
       "Centrifuge_Write_TO_T-103_DB".RequestProduct := "Centrifuge_Write_TO_T-103_DB".RouteOpened AND NOT "Centrifuge_Aux_DB"."Bool".Centrifuge.Status.FeelerRetracted;
       //************************************************Interlocks to T-104*************************************************//
       "Centrifuge_Write_TO_T-104_DB".RouteOpened := "XV-1045_DB".OS AND ("XV-3013_DB".OS OR "XV-3012_DB".OS) AND ("P-301A_DB".CF OR "P-301A_DB".CF);

       "Centrifuge_Write_TO_T-104_DB".ReqWater := "Centrifuge_DB".Status.Step = 29 AND  "Centrifuge_Write_TO_T-104_DB".RouteOpened
       AND NOT "LT-1051_DB".Alarms.HighHigh AND NOT "Centrifuge_DB".Cmds.Hold;
       //***************Valves Status***************//
       "Centrifuge_Aux_DB"."Bool".TOff := "Centrifuge_DB".Equipments.Valves."XV-1045".TurningOff OR "Centrifuge_DB".Equipments.Valves."XV-3013".TurningOff
       OR "Centrifuge_DB".Equipments.Valves."XV-3012".TurningOff OR "Centrifuge_DB".Equipments.Valves."XV-3011".TurningOff;

       //***********************************************Timers****************************************************************************//
       "Centrifuge_Aux_DB"."Bool".WaitForBucketEn := "Centrifuge_DB".Status.Step=26 AND "FT-3011_DB".SAI>1.0;
       "Centrifuge_Aux_DB"."Bool".DryingWetCakeEn := "Centrifuge_DB".Status.Step = 31  AND ("P-301A_DB".CF OR "P-301B_DB".CF) AND "FT-3012_DB".SAI < 0.1; //AND "VFD-C301R_DB".RUN_FEEDBACK
       "Centrifuge_Aux_DB"."Bool".DryingWetCake_Reset := "Centrifuge_DB".Cmds.Abort OR "Centrifuge_DB".Status.Step = 1;
       //Delay for Dry Spin Done to Finish
       "Centrifuge_Aux_DB"."Bool".DrySpinDnDelay_Enab := "Centrifuge_DB".Status.Step = 31 AND "FT-3012_DB".SAI < 0.1 AND ("P-301A_DB".CF OR "P-301B_DB".CF);
END_FUNCTION

FUNCTION "Centrifuge_SEQ_FC" : Void   // FC91, LAD
{ S7_Optimized_Access := 'TRUE' }
VERSION : 0.1
   VAR_TEMP   // added for the SCL form of the ladder/FBD networks
      _w1 : Bool;
      _w2 : Bool;
   END_VAR
BEGIN

REGION Network 2: Abort
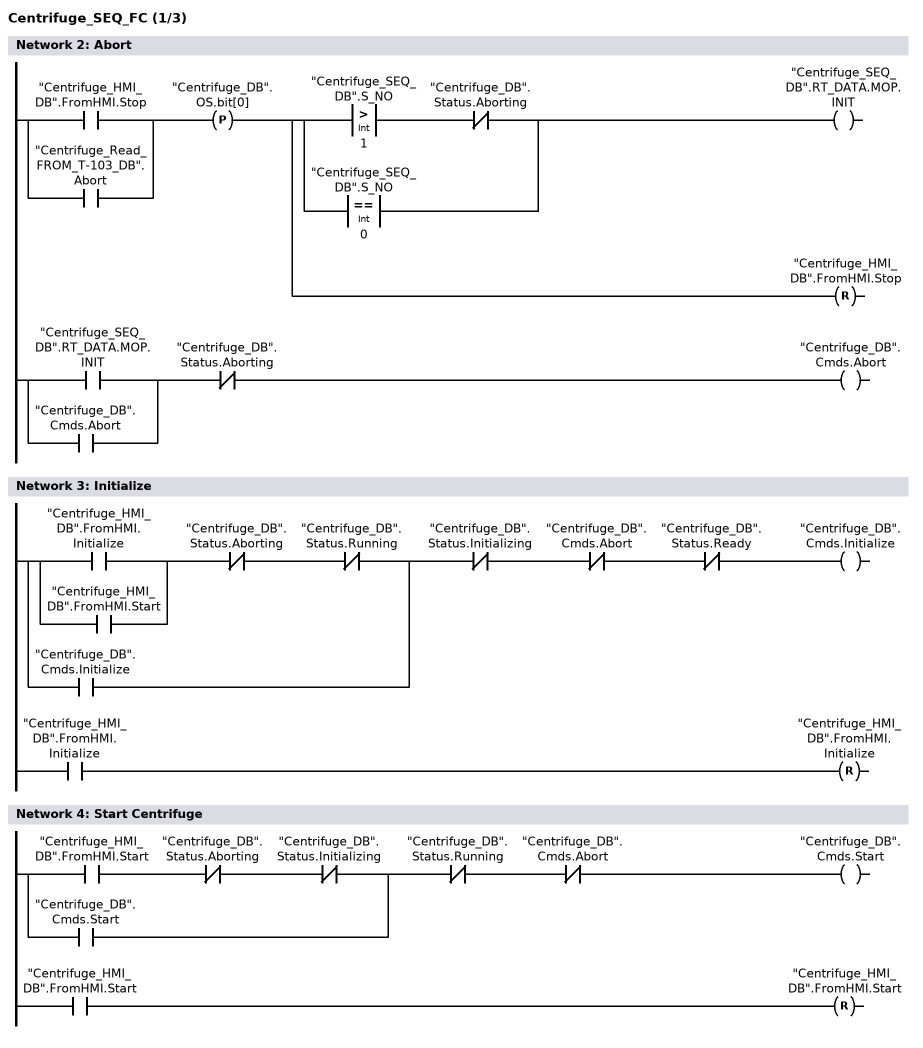
   RUNG wire#powerrail
      Contact( "Centrifuge_HMI_DB".FromHMI.Stop )
      wire#w1
      P_Trig( "Centrifuge_DB".OS.bit[0] )
      wire#w2
      { S7_Templates := "SrcType := Int" } GT_Contact(in1 := "Centrifuge_SEQ_DB".S_NO, in2 := 1)
      I_Contact( "Centrifuge_DB".Status.Aborting )
      wire#w3
      Coil( "Centrifuge_SEQ_DB".RT_DATA.MOP.INIT )
   END_RUNG
   RUNG wire#powerrail
      Contact( "Centrifuge_Read_FROM_T-103_DB".Abort )
   END_RUNG wire#w1
   RUNG wire#w2
      { S7_Templates := "SrcType := Int" } EQ_Contact(in1 := "Centrifuge_SEQ_DB".S_NO, in2 := 0)
   END_RUNG wire#w3
   RUNG wire#w2
      R_Coil( "Centrifuge_HMI_DB".FromHMI.Stop )
   END_RUNG
   RUNG wire#powerrail
      Contact( "Centrifuge_SEQ_DB".RT_DATA.MOP.INIT )
      wire#w4
      I_Contact( "Centrifuge_DB".Status.Aborting )
      Coil( "Centrifuge_DB".Cmds.Abort )
   END_RUNG
   RUNG wire#powerrail
      Contact( "Centrifuge_DB".Cmds.Abort )
   END_RUNG wire#w4
   // the same network as SCL:
   #_w1 := "Centrifuge_HMI_DB".FromHMI.Stop OR "Centrifuge_Read_FROM_T-103_DB".Abort;
   #_w2 := #_w1 AND NOT "Centrifuge_DB".OS.bit[0];   // rising edge
   "Centrifuge_DB".OS.bit[0] := #_w1;
   "Centrifuge_SEQ_DB".RT_DATA.MOP.INIT := #_w2 AND ((("Centrifuge_SEQ_DB".S_NO > 1) AND NOT "Centrifuge_DB".Status.Aborting) OR ("Centrifuge_SEQ_DB".S_NO = 0));
   IF #_w2 THEN "Centrifuge_HMI_DB".FromHMI.Stop := FALSE; END_IF;
   "Centrifuge_DB".Cmds.Abort := ("Centrifuge_SEQ_DB".RT_DATA.MOP.INIT OR "Centrifuge_DB".Cmds.Abort) AND NOT "Centrifuge_DB".Status.Aborting;
END_REGION

REGION Network 3: Initialize
   RUNG wire#powerrail
      Contact( "Centrifuge_HMI_DB".FromHMI.Initialize )
      wire#w1
      I_Contact( "Centrifuge_DB".Status.Aborting )
      I_Contact( "Centrifuge_DB".Status.Running )
      wire#w2
      I_Contact( "Centrifuge_DB".Status.Initializing )
      I_Contact( "Centrifuge_DB".Cmds.Abort )
      I_Contact( "Centrifuge_DB".Status.Ready )
      Coil( "Centrifuge_DB".Cmds.Initialize )
   END_RUNG
   RUNG wire#powerrail
      Contact( "Centrifuge_HMI_DB".FromHMI.Start )
   END_RUNG wire#w1
   RUNG wire#powerrail
      Contact( "Centrifuge_DB".Cmds.Initialize )
   END_RUNG wire#w2
   RUNG wire#powerrail
      Contact( "Centrifuge_HMI_DB".FromHMI.Initialize )
      R_Coil( "Centrifuge_HMI_DB".FromHMI.Initialize )
   END_RUNG
   // the same network as SCL:
   "Centrifuge_DB".Cmds.Initialize := ((("Centrifuge_HMI_DB".FromHMI.Initialize OR "Centrifuge_HMI_DB".FromHMI.Start) AND NOT "Centrifuge_DB".Status.Aborting AND NOT "Centrifuge_DB".Status.Running) OR "Centrifuge_DB".Cmds.Initialize) AND NOT "Centrifuge_DB".Status.Initializing AND NOT "Centrifuge_DB".Cmds.Abort AND NOT "Centrifuge_DB".Status.Ready;
   IF "Centrifuge_HMI_DB".FromHMI.Initialize THEN "Centrifuge_HMI_DB".FromHMI.Initialize := FALSE; END_IF;
END_REGION

REGION Network 4: Start Centrifuge
   RUNG wire#powerrail
      Contact( "Centrifuge_HMI_DB".FromHMI.Start )
      I_Contact( "Centrifuge_DB".Status.Aborting )
      I_Contact( "Centrifuge_DB".Status.Initializing )
      wire#w1
      I_Contact( "Centrifuge_DB".Status.Running )
      I_Contact( "Centrifuge_DB".Cmds.Abort )
      Coil( "Centrifuge_DB".Cmds.Start )
   END_RUNG
   RUNG wire#powerrail
      Contact( "Centrifuge_DB".Cmds.Start )
   END_RUNG wire#w1
   RUNG wire#powerrail
      Contact( "Centrifuge_HMI_DB".FromHMI.Start )
      R_Coil( "Centrifuge_HMI_DB".FromHMI.Start )
   END_RUNG
   // the same network as SCL:
   "Centrifuge_DB".Cmds.Start := (("Centrifuge_HMI_DB".FromHMI.Start AND NOT "Centrifuge_DB".Status.Aborting AND NOT "Centrifuge_DB".Status.Initializing) OR "Centrifuge_DB".Cmds.Start) AND NOT "Centrifuge_DB".Status.Running AND NOT "Centrifuge_DB".Cmds.Abort;
   IF "Centrifuge_HMI_DB".FromHMI.Start THEN "Centrifuge_HMI_DB".FromHMI.Start := FALSE; END_IF;
END_REGION

REGION Network 5: Procedure Selected
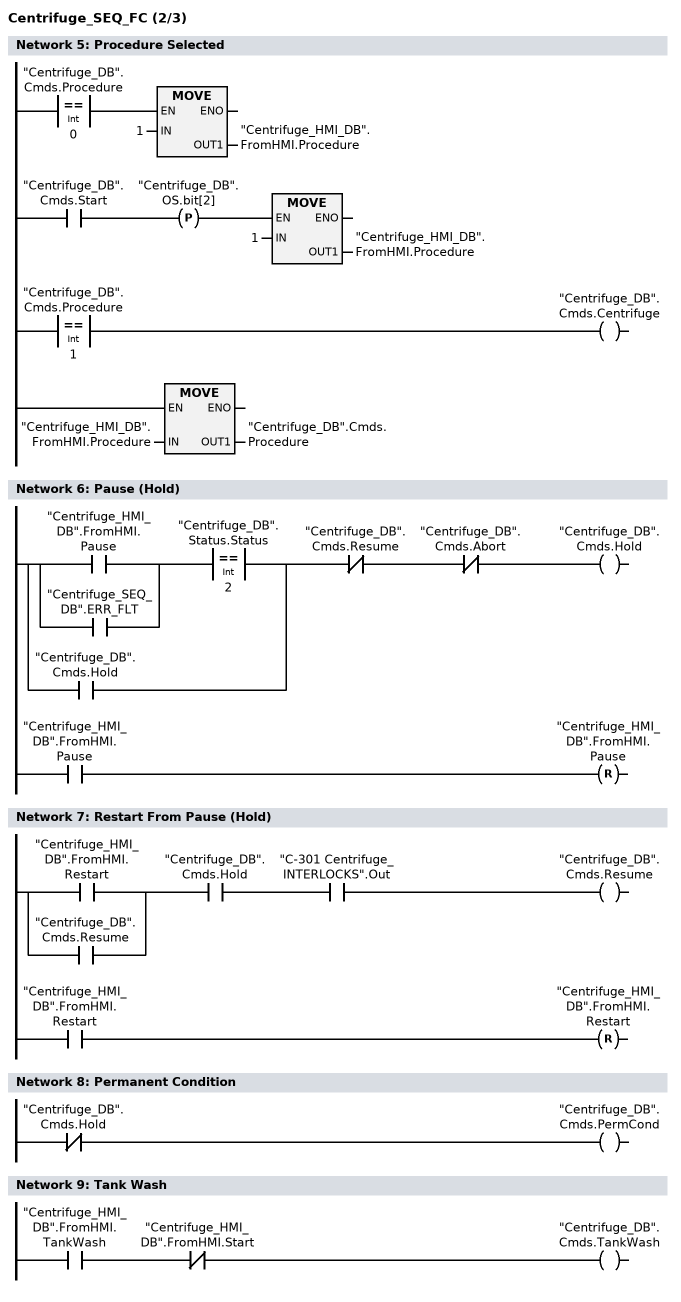
   RUNG wire#powerrail
      { S7_Templates := "SrcType := Int" } EQ_Contact(in1 := "Centrifuge_DB".Cmds.Procedure, in2 := 0)
      Move(in := 1, out1 => "Centrifuge_HMI_DB".FromHMI.Procedure)
   END_RUNG
   RUNG wire#powerrail
      Contact( "Centrifuge_DB".Cmds.Start )
      P_Trig( "Centrifuge_DB".OS.bit[2] )
      Move(in := 1, out1 => "Centrifuge_HMI_DB".FromHMI.Procedure)
   END_RUNG
   RUNG wire#powerrail
      { S7_Templates := "SrcType := Int" } EQ_Contact(in1 := "Centrifuge_DB".Cmds.Procedure, in2 := 1)
      Coil( "Centrifuge_DB".Cmds.Centrifuge )
   END_RUNG
   RUNG wire#powerrail
      Move(in := "Centrifuge_HMI_DB".FromHMI.Procedure, out1 => "Centrifuge_DB".Cmds.Procedure)
   END_RUNG
   // the same network as SCL:
   IF "Centrifuge_DB".Cmds.Procedure = 0 THEN "Centrifuge_HMI_DB".FromHMI.Procedure := 1; END_IF;
   #_w1 := "Centrifuge_DB".Cmds.Start AND NOT "Centrifuge_DB".OS.bit[2];   // rising edge
   "Centrifuge_DB".OS.bit[2] := "Centrifuge_DB".Cmds.Start;
   IF #_w1 THEN "Centrifuge_HMI_DB".FromHMI.Procedure := 1; END_IF;
   "Centrifuge_DB".Cmds.Centrifuge := "Centrifuge_DB".Cmds.Procedure = 1;
   "Centrifuge_DB".Cmds.Procedure := "Centrifuge_HMI_DB".FromHMI.Procedure;
END_REGION

REGION Network 6: Pause (Hold)
   RUNG wire#powerrail
      Contact( "Centrifuge_HMI_DB".FromHMI.Pause )
      wire#w1
      { S7_Templates := "SrcType := Int" } EQ_Contact(in1 := "Centrifuge_DB".Status.Status, in2 := 2)
      wire#w2
      I_Contact( "Centrifuge_DB".Cmds.Resume )
      I_Contact( "Centrifuge_DB".Cmds.Abort )
      Coil( "Centrifuge_DB".Cmds.Hold )
   END_RUNG
   RUNG wire#powerrail
      Contact( "Centrifuge_SEQ_DB".ERR_FLT )
   END_RUNG wire#w1
   RUNG wire#powerrail
      Contact( "Centrifuge_DB".Cmds.Hold )
   END_RUNG wire#w2
   RUNG wire#powerrail
      Contact( "Centrifuge_HMI_DB".FromHMI.Pause )
      R_Coil( "Centrifuge_HMI_DB".FromHMI.Pause )
   END_RUNG
   // the same network as SCL:
   "Centrifuge_DB".Cmds.Hold := ((("Centrifuge_HMI_DB".FromHMI.Pause OR "Centrifuge_SEQ_DB".ERR_FLT) AND ("Centrifuge_DB".Status.Status = 2)) OR "Centrifuge_DB".Cmds.Hold) AND NOT "Centrifuge_DB".Cmds.Resume AND NOT "Centrifuge_DB".Cmds.Abort;
   IF "Centrifuge_HMI_DB".FromHMI.Pause THEN "Centrifuge_HMI_DB".FromHMI.Pause := FALSE; END_IF;
END_REGION

REGION Network 7: Restart From Pause (Hold)
   RUNG wire#powerrail
      Contact( "Centrifuge_HMI_DB".FromHMI.Restart )
      wire#w1
      Contact( "Centrifuge_DB".Cmds.Hold )
      Contact( "C-301 Centrifuge_INTERLOCKS".Out )
      Coil( "Centrifuge_DB".Cmds.Resume )
   END_RUNG
   RUNG wire#powerrail
      Contact( "Centrifuge_DB".Cmds.Resume )
   END_RUNG wire#w1
   RUNG wire#powerrail
      Contact( "Centrifuge_HMI_DB".FromHMI.Restart )
      R_Coil( "Centrifuge_HMI_DB".FromHMI.Restart )
   END_RUNG
   // the same network as SCL:
   "Centrifuge_DB".Cmds.Resume := ("Centrifuge_HMI_DB".FromHMI.Restart OR "Centrifuge_DB".Cmds.Resume) AND "Centrifuge_DB".Cmds.Hold AND "C-301 Centrifuge_INTERLOCKS".Out;
   IF "Centrifuge_HMI_DB".FromHMI.Restart THEN "Centrifuge_HMI_DB".FromHMI.Restart := FALSE; END_IF;
END_REGION

REGION Network 8: Permanent Condition
   RUNG wire#powerrail
      I_Contact( "Centrifuge_DB".Cmds.Hold )
      Coil( "Centrifuge_DB".Cmds.PermCond )
   END_RUNG
   // the same network as SCL:
   "Centrifuge_DB".Cmds.PermCond := NOT "Centrifuge_DB".Cmds.Hold;
END_REGION

REGION Network 9: Tank Wash
   RUNG wire#powerrail
      Contact( "Centrifuge_HMI_DB".FromHMI.TankWash )
      I_Contact( "Centrifuge_HMI_DB".FromHMI.Start )
      Coil( "Centrifuge_DB".Cmds.TankWash )
   END_RUNG
   // the same network as SCL:
   "Centrifuge_DB".Cmds.TankWash := "Centrifuge_HMI_DB".FromHMI.TankWash AND NOT "Centrifuge_HMI_DB".FromHMI.Start;
END_REGION

REGION Network 10: Tube Wash
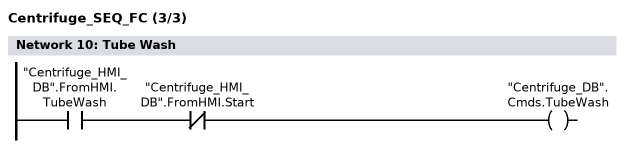
   RUNG wire#powerrail
      Contact( "Centrifuge_HMI_DB".FromHMI.TubeWash )
      I_Contact( "Centrifuge_HMI_DB".FromHMI.Start )
      Coil( "Centrifuge_DB".Cmds.TubeWash )
   END_RUNG
   // the same network as SCL:
   "Centrifuge_DB".Cmds.TubeWash := "Centrifuge_HMI_DB".FromHMI.TubeWash AND NOT "Centrifuge_HMI_DB".FromHMI.Start;
END_REGION

REGION Network 11 (SCL): Sequence Status
   IF "Centrifuge_SEQ_DB".S_NO= 1 THEN
       "Centrifuge_DB".Status.Status := 1; //Idle
   ELSIF ("Centrifuge_SEQ_DB".S_NO > 1 AND "Centrifuge_SEQ_DB".S_NO < 150) AND NOT "Centrifuge_SEQ_DB".ERR_FLT AND NOT "Centrifuge_DB".Cmds.Hold THEN
       "Centrifuge_DB".Status.Status := 2; //Running
   ELSIF "Centrifuge_SEQ_DB".S_NO >= 151 AND "Centrifuge_SEQ_DB".S_NO <= 160 AND NOT "Centrifuge_SEQ_DB".ERR_FLT THEN
       "Centrifuge_DB".Status.Status := 3; // Stopping
   ELSIF  "Centrifuge_SEQ_DB".ERR_FLT AND  ("Centrifuge_SEQ_DB".S_NO > 1 AND "Centrifuge_SEQ_DB".S_NO < 150) THEN
       "Centrifuge_DB".Status.Status := 4; // Held
   ELSIF  "Centrifuge_SEQ_DB".ERR_FLT AND  ("Centrifuge_SEQ_DB".S_NO > 1 AND "Centrifuge_SEQ_DB".S_NO < 150) AND "Centrifuge_Aux_DB"."Bool".TOff  THEN
       "Centrifuge_DB".Status.Status := 5; // Holding
   ELSE
       "Centrifuge_DB".Status.Status := 6; // Unknown
   END_IF;

   "Centrifuge_DB".Status.Running := ("Centrifuge_SEQ_DB".S_NO > 3 AND "Centrifuge_SEQ_DB".S_NO <= 150);
   "Centrifuge_DB".Status.Initializing := ("Centrifuge_SEQ_DB".S_NO >= 141 AND "Centrifuge_SEQ_DB".S_NO <= 150);

   //Enable/Disable HMI Start/Stop Button
   "Centrifuge_HMI_DB".ToHMI.EnStopButton := ("Centrifuge_DB".Status.Status > 1) OR "Centrifuge_DB".Status.Step = 0; //Enable HMI Stop Button
   "Centrifuge_HMI_DB".ToHMI.EnStartButton := "Centrifuge_DB".Status.Status = 1; //Idle
   "Centrifuge_HMI_DB".ToHMI.EnPauseButton := "Centrifuge_DB".Status.Status = 2; //Enable Pause Button
   "Centrifuge_HMI_DB".ToHMI.EnRestartButton :=  "Centrifuge_DB".Status.Status = 4; //Enable Restart Button

   //****Interlock Activated
   "Centrifuge_HMI_DB".ToHMI.InterlockActivated := "C-301 Centrifuge_INTERLOCKS".Out;
END_REGION

REGION Network 12 (SCL): Sequence Step
   "Centrifuge_DB".Status.Step := "Centrifuge_SEQ_DB".S_NO;
END_REGION

REGION Network 13 (SCL): Sequence state (Procedure running)
   IF "Centrifuge_SEQ_DB".S_NO = 3 OR "Centrifuge_SEQ_DB".S_NO = 4 THEN
       "Centrifuge_DB".Status.State := 1; //Ready
   ELSIF "Centrifuge_SEQ_DB".S_NO >= 21 AND "Centrifuge_SEQ_DB".S_NO <= 60 THEN
       "Centrifuge_DB".Status.State := 2; //Mixing 
   ELSIF "Centrifuge_SEQ_DB".S_NO >= 61 AND "Centrifuge_SEQ_DB".S_NO <= 80 THEN
       "Centrifuge_DB".Status.State := 3; //Pouring
   ELSIF "Centrifuge_SEQ_DB".S_NO >= 141 AND "Centrifuge_SEQ_DB".S_NO <= 150 THEN
       "Centrifuge_DB".Status.State := 4; //Initializing
   ELSIF "Centrifuge_SEQ_DB".S_NO >= 151 AND "Centrifuge_SEQ_DB".S_NO <= 160 THEN
       "Centrifuge_DB".Status.State := 5; //Aborting
   ELSE
       "Centrifuge_DB".Status.State := 0;
   END_IF;
END_REGION

REGION Network 14: Sequence State
END_REGION
END_FUNCTION

FUNCTION "Centrifuge_AuxOutputs_FC" : Void   // FC109, LAD
{ S7_Optimized_Access := 'TRUE' }
VERSION : 0.1
   VAR_TEMP   // added for the SCL form of the ladder/FBD networks
      _w1 : Bool;
   END_VAR
BEGIN

REGION Network 1: Centrifuge Start Command
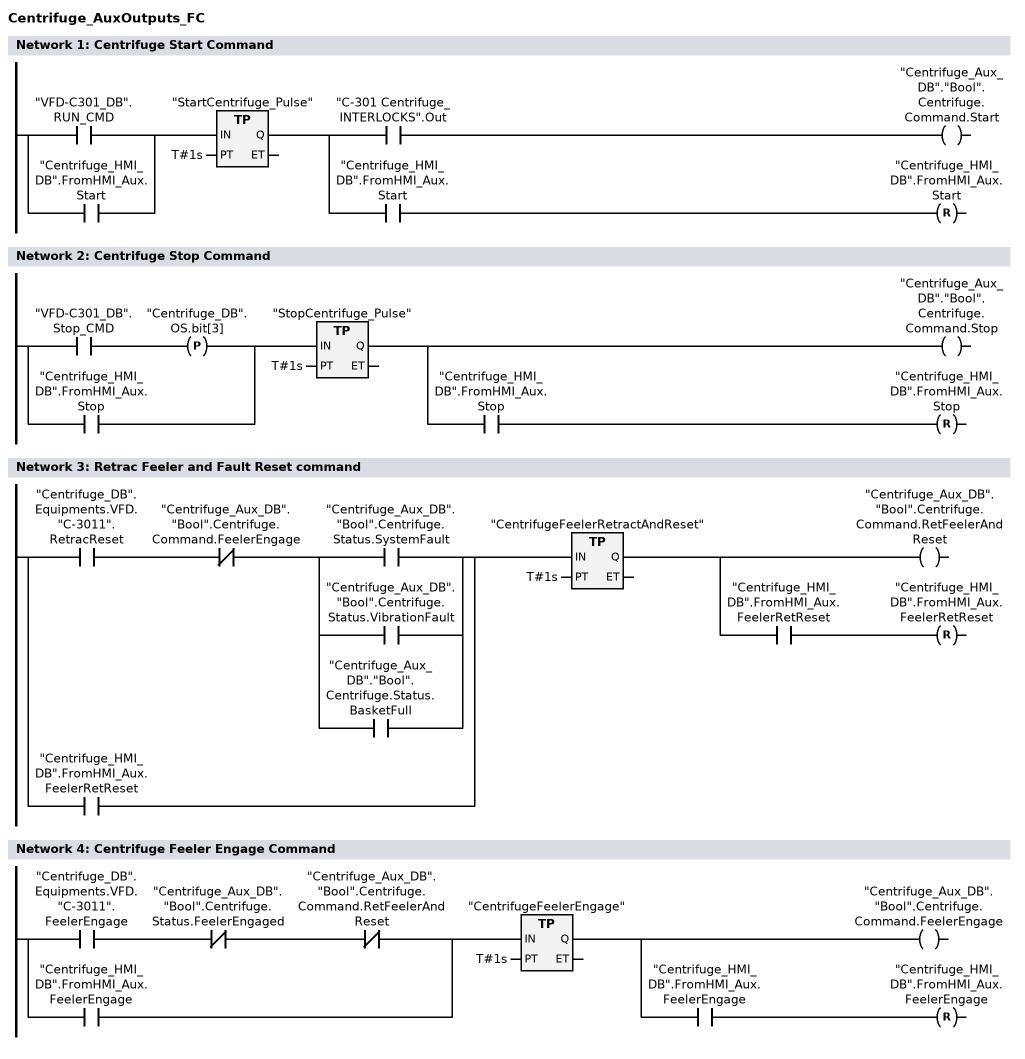
   "StartCentrifuge_Pulse".TP(IN := "VFD-C301_DB".RUN_CMD OR "Centrifuge_HMI_DB".FromHMI_Aux.Start, PT := T#1s);
   "Centrifuge_Aux_DB"."Bool".Centrifuge.Command.Start := "StartCentrifuge_Pulse".Q AND "C-301 Centrifuge_INTERLOCKS".Out;
   IF "StartCentrifuge_Pulse".Q AND "Centrifuge_HMI_DB".FromHMI_Aux.Start THEN
       "Centrifuge_HMI_DB".FromHMI_Aux.Start := FALSE;
   END_IF;
END_REGION

REGION Network 2: Centrifuge Stop Command
   #_w1 := "VFD-C301_DB".Stop_CMD AND NOT "Centrifuge_DB".OS.bit[3];   // rising edge
   "Centrifuge_DB".OS.bit[3] := "VFD-C301_DB".Stop_CMD;
   "StopCentrifuge_Pulse".TP(IN := #_w1 OR "Centrifuge_HMI_DB".FromHMI_Aux.Stop, PT := T#1s);
   "Centrifuge_Aux_DB"."Bool".Centrifuge.Command.Stop := "StopCentrifuge_Pulse".Q;
   IF "StopCentrifuge_Pulse".Q AND "Centrifuge_HMI_DB".FromHMI_Aux.Stop THEN
       "Centrifuge_HMI_DB".FromHMI_Aux.Stop := FALSE;
   END_IF;
END_REGION

REGION Network 3: Retrac Feeler and Fault Reset command
   "CentrifugeFeelerRetractAndReset".TP(IN := ("Centrifuge_DB".Equipments.VFD."C-3011".RetracReset AND NOT "Centrifuge_Aux_DB"."Bool".Centrifuge.Command.FeelerEngage AND ("Centrifuge_Aux_DB"."Bool".Centrifuge.Status.SystemFault OR "Centrifuge_Aux_DB"."Bool".Centrifuge.Status.VibrationFault OR "Centrifuge_Aux_DB"."Bool".Centrifuge.Status.BasketFull)) OR "Centrifuge_HMI_DB".FromHMI_Aux.FeelerRetReset,
                           PT := T#1s);
   "Centrifuge_Aux_DB"."Bool".Centrifuge.Command.RetFeelerAndReset := "CentrifugeFeelerRetractAndReset".Q;
   IF "CentrifugeFeelerRetractAndReset".Q AND "Centrifuge_HMI_DB".FromHMI_Aux.FeelerRetReset THEN
       "Centrifuge_HMI_DB".FromHMI_Aux.FeelerRetReset := FALSE;
   END_IF;
END_REGION

REGION Network 4: Centrifuge Feeler Engage Command
   "CentrifugeFeelerEngage".TP(IN := ("Centrifuge_DB".Equipments.VFD."C-3011".FeelerEngage AND NOT "Centrifuge_Aux_DB"."Bool".Centrifuge.Status.FeelerEngaged AND NOT "Centrifuge_Aux_DB"."Bool".Centrifuge.Command.RetFeelerAndReset) OR "Centrifuge_HMI_DB".FromHMI_Aux.FeelerEngage,
                           PT := T#1s);
   "Centrifuge_Aux_DB"."Bool".Centrifuge.Command.FeelerEngage := "CentrifugeFeelerEngage".Q;
   IF "CentrifugeFeelerEngage".Q AND "Centrifuge_HMI_DB".FromHMI_Aux.FeelerEngage THEN
       "Centrifuge_HMI_DB".FromHMI_Aux.FeelerEngage := FALSE;
   END_IF;
END_REGION
END_FUNCTION

FUNCTION "Centrifuge_Transitions_FC" : Void   // FC110, SCL
{ S7_Optimized_Access := 'TRUE' }
VERSION : 0.1
BEGIN
   //*************************Transitions********************************
   //Initials Done
   "Centrifuge_DB".Transitions.InitialsDone := "XV-1045_DB".CS AND "XV-3013_DB".CS AND "XV-3012_DB".CS AND "FV-3011_DB".CMD = 0.0
   AND NOT "P-301A_DB".CF AND NOT "P-301B_DB".CF AND "FT-3012_Totalizer_DB".Total = 0.0 AND "FT-3011_Totalizer_DB".Total = 0.0
   AND "FT-1045_Totalizer_DB".Total = 0.0 AND NOT "Centrifuge_Aux_DB"."Bool".Centrifuge.Command.RetFeelerAndReset;

   //Ready to Run
   "Centrifuge_DB".Transitions.ReadytoRun :=  "Centrifuge_Aux_DB"."Bool".Centrifuge.Status.FeelerEngaged
   AND NOT "Centrifuge_Aux_DB"."Bool".Centrifuge.Status.SystemFault AND NOT "Centrifuge_Aux_DB"."Bool".Centrifuge.Status.VibrationFault
   AND "Centrifuge_Aux_DB"."Bool".Centrifuge.Status.CoverLocked AND NOT "Centrifuge_Aux_DB"."Bool".Centrifuge.Command.FeelerEngage;

   //Basket Full
   "Centrifuge_DB".Transitions.BasketFull := "Centrifuge_Aux_DB"."Bool".Centrifuge.Status.BasketFull;
END_FUNCTION

// folder: State MACHINE/3)Centrifuge/Centrifuge <---> T-103

FUNCTION "Centrifuge_Signals_FROM_T-103" : Void   // FC68, LAD
{ S7_Optimized_Access := 'TRUE' }
VERSION : 0.1
BEGIN

REGION Network 1: Started Sequence
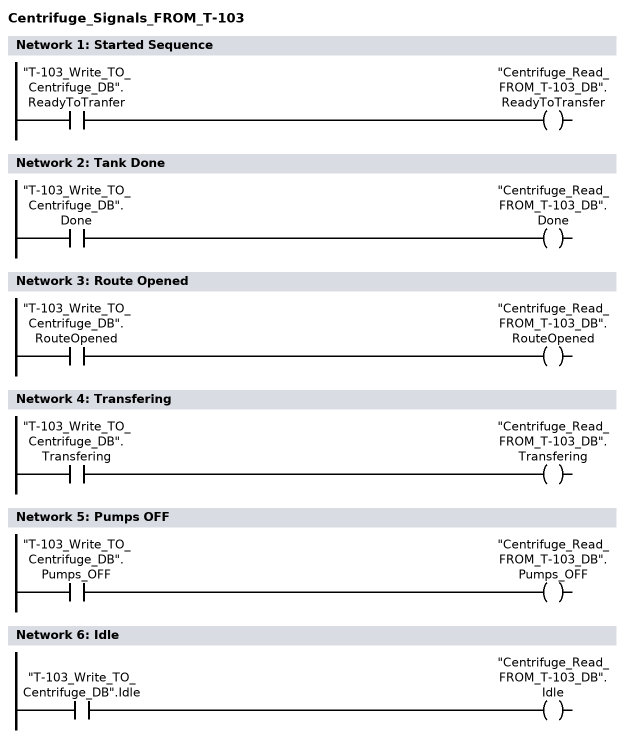
   RUNG wire#powerrail
      Contact( "T-103_Write_TO_Centrifuge_DB".ReadyToTranfer )
      Coil( "Centrifuge_Read_FROM_T-103_DB".ReadyToTransfer )
   END_RUNG
   // the same network as SCL:
   "Centrifuge_Read_FROM_T-103_DB".ReadyToTransfer := "T-103_Write_TO_Centrifuge_DB".ReadyToTranfer;
END_REGION

REGION Network 2: Tank Done
   RUNG wire#powerrail
      Contact( "T-103_Write_TO_Centrifuge_DB".Done )
      Coil( "Centrifuge_Read_FROM_T-103_DB".Done )
   END_RUNG
   // the same network as SCL:
   "Centrifuge_Read_FROM_T-103_DB".Done := "T-103_Write_TO_Centrifuge_DB".Done;
END_REGION

REGION Network 3: Route Opened
   RUNG wire#powerrail
      Contact( "T-103_Write_TO_Centrifuge_DB".RouteOpened )
      Coil( "Centrifuge_Read_FROM_T-103_DB".RouteOpened )
   END_RUNG
   // the same network as SCL:
   "Centrifuge_Read_FROM_T-103_DB".RouteOpened := "T-103_Write_TO_Centrifuge_DB".RouteOpened;
END_REGION

REGION Network 4: Transfering
   RUNG wire#powerrail
      Contact( "T-103_Write_TO_Centrifuge_DB".Transfering )
      Coil( "Centrifuge_Read_FROM_T-103_DB".Transfering )
   END_RUNG
   // the same network as SCL:
   "Centrifuge_Read_FROM_T-103_DB".Transfering := "T-103_Write_TO_Centrifuge_DB".Transfering;
END_REGION

REGION Network 5: Pumps OFF
   RUNG wire#powerrail
      Contact( "T-103_Write_TO_Centrifuge_DB".Pumps_OFF )
      Coil( "Centrifuge_Read_FROM_T-103_DB".Pumps_OFF )
   END_RUNG
   // the same network as SCL:
   "Centrifuge_Read_FROM_T-103_DB".Pumps_OFF := "T-103_Write_TO_Centrifuge_DB".Pumps_OFF;
END_REGION

REGION Network 6: Idle
   RUNG wire#powerrail
      Contact( "T-103_Write_TO_Centrifuge_DB".Idle )
      Coil( "Centrifuge_Read_FROM_T-103_DB".Idle )
   END_RUNG
   // the same network as SCL:
   "Centrifuge_Read_FROM_T-103_DB".Idle := "T-103_Write_TO_Centrifuge_DB".Idle;
END_REGION
END_FUNCTION

// folder: State MACHINE/3)Centrifuge/Centrifuge <---> T-104

FUNCTION "Centrifuge_Signals_FROM_T-104" : Void   // FC67, LAD
{ S7_Optimized_Access := 'TRUE' }
VERSION : 0.1
BEGIN

REGION Network 1: Ready
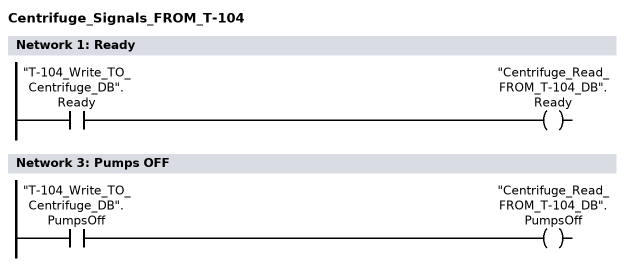
   RUNG wire#powerrail
      Contact( "T-104_Write_TO_Centrifuge_DB".Ready )
      Coil( "Centrifuge_Read_FROM_T-104_DB".Ready )
   END_RUNG
   // the same network as SCL:
   "Centrifuge_Read_FROM_T-104_DB".Ready := "T-104_Write_TO_Centrifuge_DB".Ready;
END_REGION

REGION Network 2: Route Opened
END_REGION

REGION Network 3: Pumps OFF
   RUNG wire#powerrail
      Contact( "T-104_Write_TO_Centrifuge_DB".PumpsOff )
      Coil( "Centrifuge_Read_FROM_T-104_DB".PumpsOff )
   END_RUNG
   // the same network as SCL:
   "Centrifuge_Read_FROM_T-104_DB".PumpsOff := "T-104_Write_TO_Centrifuge_DB".PumpsOff;
END_REGION
END_FUNCTION

// folder: State MACHINE/4)Calcination

FUNCTION "Monitor_SEQ_FC" : Void   // FC28, LAD
TITLE = FC to call User Functions
{ S7_Optimized_Access := 'TRUE' }
AUTHOR : JL
VERSION : 0.1
BEGIN

REGION Network 1: Moving Furnace temperature to the monitor block
   // Thermocouples:
   // "TT-401A_DB".SAI
   // "TT-401B_DB".SAI
   // "TT-401C_DB".SAI
   // "TT-401C_DB".SAI
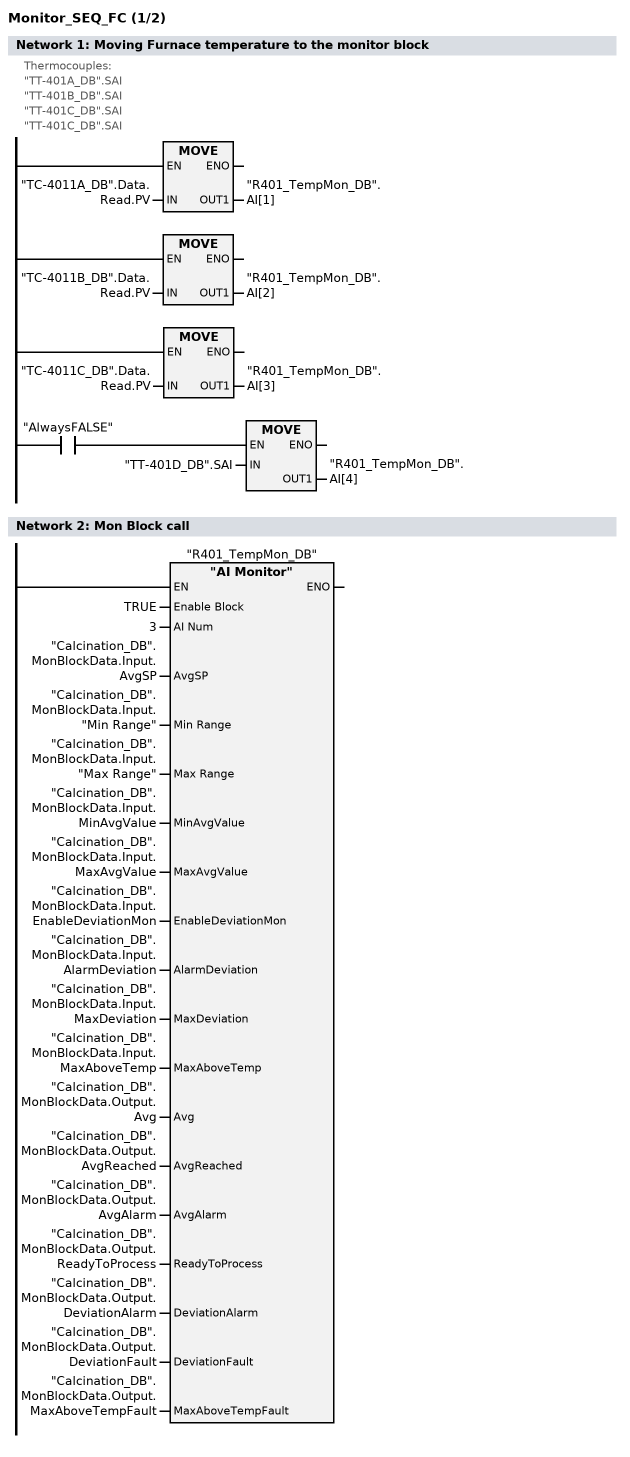
   RUNG wire#powerrail
      Move(in := "TC-4011A_DB".Data.Read.PV, out1 => "R401_TempMon_DB".AI[1])
   END_RUNG
   RUNG wire#powerrail
      Move(in := "TC-4011B_DB".Data.Read.PV, out1 => "R401_TempMon_DB".AI[2])
   END_RUNG
   RUNG wire#powerrail
      Move(in := "TC-4011C_DB".Data.Read.PV, out1 => "R401_TempMon_DB".AI[3])
   END_RUNG
   RUNG wire#powerrail
      Contact( "AlwaysFALSE" )
      Move(in := "TT-401D_DB".SAI, out1 => "R401_TempMon_DB".AI[4])
   END_RUNG
   // the same network as SCL:
   "R401_TempMon_DB".AI[1] := "TC-4011A_DB".Data.Read.PV;
   "R401_TempMon_DB".AI[2] := "TC-4011B_DB".Data.Read.PV;
   "R401_TempMon_DB".AI[3] := "TC-4011C_DB".Data.Read.PV;
   IF "AlwaysFALSE" THEN "R401_TempMon_DB".AI[4] := "TT-401D_DB".SAI; END_IF;
END_REGION

REGION Network 2: Mon Block call
   RUNG wire#powerrail
      "R401_TempMon_DB"("Enable Block" := TRUE, "AI Num" := 3, AvgSP := "Calcination_DB".MonBlockData.Input.AvgSP, "Min Range" := "Calcination_DB".MonBlockData.Input."Min Range", "Max Range" := "Calcination_DB".MonBlockData.Input."Max Range", MinAvgValue := "Calcination_DB".MonBlockData.Input.MinAvgValue, MaxAvgValue := "Calcination_DB".MonBlockData.Input.MaxAvgValue, EnableDeviationMon := "Calcination_DB".MonBlockData.Input.EnableDeviationMon, AlarmDeviation := "Calcination_DB".MonBlockData.Input.AlarmDeviation, MaxDeviation := "Calcination_DB".MonBlockData.Input.MaxDeviation, MaxAboveTemp := "Calcination_DB".MonBlockData.Input.MaxAboveTemp, Avg := "Calcination_DB".MonBlockData.Output.Avg, AvgReached := "Calcination_DB".MonBlockData.Output.AvgReached, AvgAlarm := "Calcination_DB".MonBlockData.Output.AvgAlarm, ReadyToProcess := "Calcination_DB".MonBlockData.Output.ReadyToProcess, DeviationAlarm := "Calcination_DB".MonBlockData.Output.DeviationAlarm, DeviationFault := "Calcination_DB".MonBlockData.Output.DeviationFault, MaxAboveTempFault := "Calcination_DB".MonBlockData.Output.MaxAboveTempFault)
   END_RUNG
   // the same network as SCL:
   "R401_TempMon_DB"("Enable Block" := TRUE,   // "AI Monitor"
                     "AI Num" := 3,
                     AvgSP := "Calcination_DB".MonBlockData.Input.AvgSP,
                     "Min Range" := "Calcination_DB".MonBlockData.Input."Min Range",
                     "Max Range" := "Calcination_DB".MonBlockData.Input."Max Range",
                     MinAvgValue := "Calcination_DB".MonBlockData.Input.MinAvgValue,
                     MaxAvgValue := "Calcination_DB".MonBlockData.Input.MaxAvgValue,
                     EnableDeviationMon := "Calcination_DB".MonBlockData.Input.EnableDeviationMon,
                     AlarmDeviation := "Calcination_DB".MonBlockData.Input.AlarmDeviation,
                     MaxDeviation := "Calcination_DB".MonBlockData.Input.MaxDeviation,
                     MaxAboveTemp := "Calcination_DB".MonBlockData.Input.MaxAboveTemp,
                     Avg := "Calcination_DB".MonBlockData.Output.Avg,
                     AvgReached := "Calcination_DB".MonBlockData.Output.AvgReached,
                     AvgAlarm := "Calcination_DB".MonBlockData.Output.AvgAlarm,
                     ReadyToProcess := "Calcination_DB".MonBlockData.Output.ReadyToProcess,
                     DeviationAlarm := "Calcination_DB".MonBlockData.Output.DeviationAlarm,
                     DeviationFault := "Calcination_DB".MonBlockData.Output.DeviationFault,
                     MaxAboveTempFault := "Calcination_DB".MonBlockData.Output.MaxAboveTempFault);
END_REGION

REGION Network 3: AIs Monitor new block
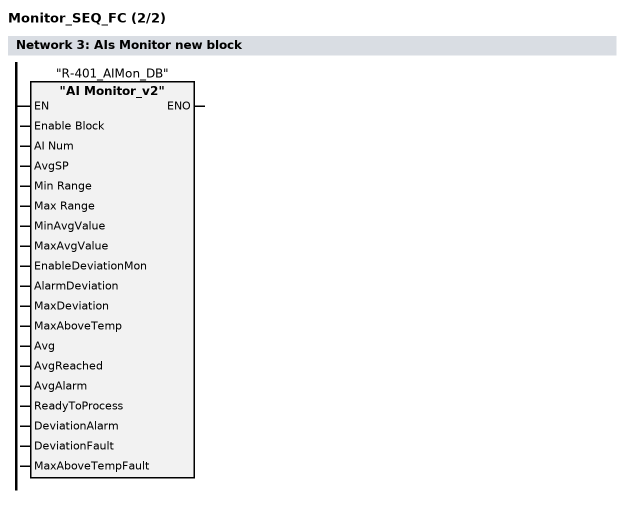
   RUNG wire#powerrail
      "R-401_AIMon_DB"("Enable Block" :=, "AI Num" :=, AvgSP :=, "Min Range" :=, "Max Range" :=, MinAvgValue :=, MaxAvgValue :=, EnableDeviationMon :=, AlarmDeviation :=, MaxDeviation :=, MaxAboveTemp :=, Avg :=, AvgReached :=, AvgAlarm :=, ReadyToProcess :=, DeviationAlarm :=, DeviationFault :=, MaxAboveTempFault :=)
   END_RUNG
   // the same network as SCL:
   "R-401_AIMon_DB"();   // "AI Monitor_v2"
END_REGION
END_FUNCTION

FUNCTION "Alarms" : Void   // FC29, LAD
{ S7_Optimized_Access := 'TRUE' }
VERSION : 0.1
   VAR_TEMP
      EurothermCommFault : Bool;
   END_VAR
BEGIN

REGION Network 1 (SCL): MFC Communication Fault (Pressure Control)
   "R-402_Aux_DB".Timer.Alarms.MFC_Cmms1.TON(IN := "MFC-4011_MB_R_DB".MB_CLIENT_Instance.DONE,
                                                    PT := T#10s);
   "R-402_Aux_DB".Timer.Alarms.MFC_Cmms2.TON(IN := NOT "MFC-4011_MB_R_DB".MB_CLIENT_Instance.DONE,
                                             PT := T#10s);

   "MFC-4011_DB_MB".Data.Status.CommFault := "R-402_Aux_DB".Timer.Alarms.MFC_Cmms1.Q OR "R-402_Aux_DB".Timer.Alarms.MFC_Cmms2.Q;
END_REGION

REGION Network 2 (SCL): Eurotherm Controllers Alarm Communications(Temperature Controllers)
   //TC-4011A Communication monitoring
   "R-402_Aux_DB".Timer.Alarms."TC-4011A_Cmms1".TON(IN := "TC-4011A_R1".MB_CLIENT_Instance.DONE,
                                                    PT := T#10s);
   "R-402_Aux_DB".Timer.Alarms."TC-4011A_Cmms2".TON(IN := NOT "TC-4011A_R1".MB_CLIENT_Instance.DONE,
                                                    PT := T#10s);
   "R-402_Aux_DB".Timer.Alarms."TC-4011B_Cmms1".TON(IN := "TC-4011B_R1".MB_CLIENT_Instance.DONE,
                                                    PT := T#10s);
   "R-402_Aux_DB".Timer.Alarms."TC-4011B_Cmms2".TON(IN := NOT "TC-4011B_R1".MB_CLIENT_Instance.DONE,
                                                    PT := T#10s);
   "R-402_Aux_DB".Timer.Alarms."TC-4011C_Cmms1".TON(IN := "TC-4011C_R1".MB_CLIENT_Instance.DONE,
                                                    PT := T#10s);
   "R-402_Aux_DB".Timer.Alarms."TC-4011C_Cmms2".TON(IN := NOT "TC-4011C_R1".MB_CLIENT_Instance.DONE,
                                                    PT := T#10s);

   "R-402_Aux_DB"."Bool".EurothermStatus."4011A_Connected" := NOT( "R-402_Aux_DB".Timer.Alarms."TC-4011A_Cmms1".Q OR "R-402_Aux_DB".Timer.Alarms."TC-4011A_Cmms2".Q);
   "R-402_Aux_DB"."Bool".EurothermStatus."4011B_Connected" := NOT ("R-402_Aux_DB".Timer.Alarms."TC-4011B_Cmms1".Q OR "R-402_Aux_DB".Timer.Alarms."TC-4011B_Cmms2".Q);
   "R-402_Aux_DB"."Bool".EurothermStatus."4011C_Connected" := NOT ("R-402_Aux_DB".Timer.Alarms."TC-4011C_Cmms1".Q OR "R-402_Aux_DB".Timer.Alarms."TC-4011C_Cmms2".Q);

   #EurothermCommFault := NOT ("R-402_Aux_DB"."Bool".EurothermStatus."4011A_Connected" AND "R-402_Aux_DB"."Bool".EurothermStatus."4011B_Connected"
   AND "R-402_Aux_DB"."Bool".EurothermStatus."4011C_Connected");
END_REGION

REGION Network 3
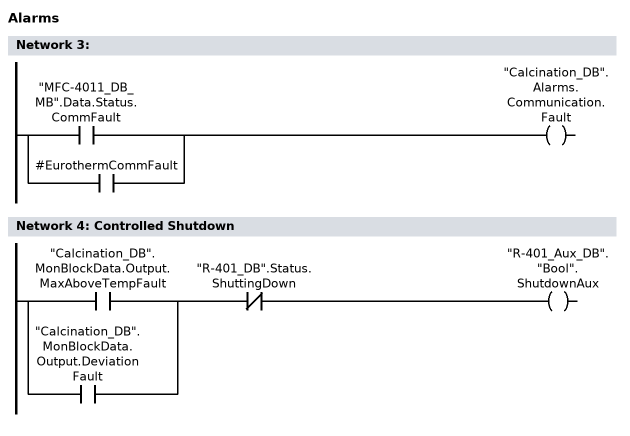
   RUNG wire#powerrail
      Contact( "MFC-4011_DB_MB".Data.Status.CommFault )
      wire#w1
      Coil( "Calcination_DB".Alarms.Communication.Fault )
   END_RUNG
   RUNG wire#powerrail
      Contact( #EurothermCommFault )
   END_RUNG wire#w1
   // the same network as SCL:
   "Calcination_DB".Alarms.Communication.Fault := "MFC-4011_DB_MB".Data.Status.CommFault OR #EurothermCommFault;
END_REGION

REGION Network 4: Controlled Shutdown
   RUNG wire#powerrail
      Contact( "Calcination_DB".MonBlockData.Output.MaxAboveTempFault )
      wire#w1
      I_Contact( "R-401_DB".Status.ShuttingDown )
      Coil( "R-401_Aux_DB"."Bool".ShutdownAux )
   END_RUNG
   RUNG wire#powerrail
      Contact( "Calcination_DB".MonBlockData.Output.DeviationFault )
   END_RUNG wire#w1
   // the same network as SCL:
   "R-401_Aux_DB"."Bool".ShutdownAux := ("Calcination_DB".MonBlockData.Output.MaxAboveTempFault OR "Calcination_DB".MonBlockData.Output.DeviationFault) AND NOT "R-401_DB".Status.ShuttingDown;
END_REGION
END_FUNCTION

// folder: State MACHINE/4)Calcination/Reactor R-401

